(* Logix 5000 project; controller PLC_MCC1300_75F1 vendor 1 type 14 code 166 rev 32.11; software revision 32.04; part 73 of 83 *)
(* tags used below, declared in another part *)
   GP_OB_InitializeMain : GP_OB_Initialize;
   GP_RampSpace : GP_RampSpace;
   GP_ScadaPlate : GP_ScadaPlate;
   Gp_SpaceConvUtilities_V1 : GP_SpaceConvUtilities_V1;
   M351 : MAC_Conveyor;
   M351_Data : UDT_Convoy_SL;
   M351_SpaceConv_Utilities : SpaceConv_Utilities;
   M352 : MAC_Conveyor;
   M352_ALM : MAC_Conveyor_ALM;
   M352_Data : UDT_Convoy_SL;
   M352_DeletePlate : BOOL;
   M352_HMR : MAC_Conveyor_HMR;
   M352_HMW : MAC_Conveyor_HMW;
   M352_Input_xPbDeleteGlass : BOOL;
   M352_Input_xPbFanOff : BOOL;   // W204SB3/A. Fan off
   M352_Input_xPbSendToCullet : BOOL;   // W204SB2. Send to cullet
   M352_M1_DR : AXIS_CIP_DRIVE;
   M352_ONS_SetResetPresence : BOOL;
   M352_SpaceConv_Utilities : SpaceConv_Utilities;
   O : INT[128];
   TMP_dConveyorNumberForZoneCleaning : DINT;
   TMP_dDecelerationPositionEndConveyor : DINT;
   TMP_dOffsetLoadUnload_cmm : DINT;
   TMP_SendToCullet : BOOL;
   TMP_x : BOOL;
   TMP_xConveyorInvolvedInCleaning : BOOL;
   TMP_xConveyorOfStartCleaning : BOOL;
   TMP_xEnableLoadUnload : BOOL;
   TMP_xEnableZoneCleaning : BOOL;
   xAlwaysOFF : BOOL;
   xAlwaysON : BOOL;
   xSampleTablePedal : BOOL;
   Z900 : MAC_Zone;
   Z900_HMI_rgtPlateScada_Internal : HMI_LiteData[5,2,7];
   Z900_HMW : MAC_Zone_HMW;
(* MainProgram, continued *)

ROUTINE M352_Alarm   (* ladder *)
   0: NOP();
   // Reset Alarm
   1: XIC(Z900.tmON_ResetAlarm.DN)FLL(0,M352_ALM,1);
   2: XIC(Z900.ST_xEnableControlError)XIC(xAlwaysOFF)XIO(M352.INPUT_xProtectionMotor_M1)OTL(M352_ALM.rgxStoppingFault_M[0].0);
   3: XIC(Z900.ST_xEnableControlError)XIC(M352.INPUT_xDriveError_M1)OTL(M352_ALM.rgxStoppingFault_M[0].1);
   4: XIC(Z900.ST_xEnableControlError)XIO(M352.INPUT_xDriveError_M1)[XIC(M352.OUTPUT_xRun_M1) ,XIC(M352.OUTPUT_xReverse_M1) ,XIC(M352.OUTPUT_xPositioning_M1) ]XIO(M352.INPUT_xDriveFeedback_M1)[XIO(M352.tmON_FeedbackTimeOut_M1.DN) TON(M352.tmON_FeedbackTimeOut_M1,?,?) ,XIC(M352.tmON_FeedbackTimeOut_M1.DN) OTL(M352_ALM.rgxStoppingFault_M[0].2) ];
   5: XIC(Z900.ST_xEnableControlError)XIC(xAlwaysOFF)XIO(M352.INPUT_xLocalSafetySwitch_M1)OTL(M352_ALM.rgxStoppingFault_M[0].3);
   6: XIC(Z900.ST_xEnableControlError)XIO(M352.INPUT_xMotorThermalProbe_M1)OTL(M352_ALM.rgxStoppingFault_M[0].4);
   7: XIC(Z900.ST_xEnableControlError)XIC(xAlwaysOFF)XIO(M352.INPUT_xBrakingResistor_M1)OTL(M352_ALM.rgxStoppingFault_M[0].5);
   8: XIC(Z900.ST_xEnableControlError)XIC(xAlwaysOFF)[XIC(M352.INPUT_xDriveInhibit_M1) ,XIC(M352.OUTPUT_xDriveEnable_M1) XIO(M352.INPUT_xDriveReady_M1) ]OTL(M352_ALM.rgxStoppingFault_M[0].6);
   9: XIC(M352.ST_xEnableControlError)XIC(xAlwaysOFF)XIC(M352.PH_x.23)NEQ(M352_SpaceConv_Utilities.CONST_dSyncMode,0)[XIO(M352.ST_xPlateSynchronized) OTL(M352_ALM.rgxWarning[0].0) ,XIC(M352.ST_xPlateSynchronized) OTU(M352_ALM.rgxWarning[0].0) ];
   10: XIC(M352.ST_xEnableControlError)XIC(xAlwaysOFF)XIC(M352.PH_x.23)[XIC(M352_Data.tFlag.tConveyor.xReqStop) ,XIC(M352_Data.tFlag.tConveyor.xBypassReqEndStop) ]OTL(M352_ALM.rgxWarning[0].1);
   // #####_CUMULATIVE ALARM_#####
   11: NOP();
   12: [NEQ(M352_ALM.rgxStoppingFault[0],0) ,NEQ(M352_ALM.rgxStoppingFault_M[0],0) ,NEQ(M352_ALM.rgxStoppingFault_M[1],0) ]OTE(M352.ST_xStopMachineFault);
   13: [NEQ(M352_ALM.rgxFault[0],0) ,NEQ(M352_ALM.rgxFault_M[0],0) ,NEQ(M352_ALM.rgxFault_M[1],0) ]OTE(M352.ST_xStopNextCycleFault);
END_ROUTINE

ROUTINE M352_Logic   (* ladder *)
   // #####_COSTANTS_#####
   0: [MOV(6010,TMP_dConveyorNumberForZoneCleaning) MOV(50000,TMP_dOffsetLoadUnload_cmm) MOV(500,M352_SpaceConv_Utilities.CONST_dPresetFeedbackTime_ms) OTU(TMP_xEnableLoadUnload) OTU(TMP_xEnableZoneCleaning) MOV(500000,M352_SpaceConv_Utilities.CONST_dConveyorLength_cmm) MOV(400000,M352_SpaceConv_Utilities.CONST_dConveyorWidth_cmm) SUB(M352_SpaceConv_Utilities.CONST_dConveyorLength_cmm,M352.AUX_dAccSpace_cmm,M352.AUX_dPresetStopLoad_cmm) ADD(M352_SpaceConv_Utilities.CONST_dConveyorLength_cmm,M352.AUX_dDecSpace_cmm,M352.AUX_dPresetStopUnload_cmm) MOV(1.2,M352_SpaceConv_Utilities.CONST_rAcceleration_ms2) MOV(1.2,M352_SpaceConv_Utilities.CONST_rDeceleration_ms2) ,[MOV(1,M352_SpaceConv_Utilities.CONST_dSyncMode) ,MOV(0,M352_SpaceConv_Utilities.CONST_dSyncroPhPosition_cmm) ,MOV(200000,M352_SpaceConv_Utilities.CONST_dSyncroPhWindow_cmm) ] ];
   // #####_MATCH_#####
   1: NOP();
   // Conveyor Cleaning
   2: XIC(TMP_xEnableZoneCleaning)XIC(Z900.ST_xCleaningAccepted)GRT(Z900_HMW.dCleaningSelection,0)[EQU(Z900_HMW.dCleaningSelection,TMP_dConveyorNumberForZoneCleaning) OTE(TMP_xConveyorOfStartCleaning) ,GEQ(Z900_HMW.dCleaningSelection,TMP_dConveyorNumberForZoneCleaning) OTE(TMP_xConveyorInvolvedInCleaning) ];
   // Enable control error
   3: XIC(Z900.ST_xEnableControlError)OTE(M352.ST_xEnableControlError);
   // Mode 7 - Offsett for load/unload Simultaney
   4: XIC(M352.PH_x.8)MOV(M352.AUX_dPresetStopLoad_cmm,M352_SpaceConv_Utilities.ST_dStopLoadForseen_cmm)MOV(TMP_dOffsetLoadUnload_cmm,M352_SpaceConv_Utilities.CONF_MD7_dOffset_cmm)GP_SpaceConvUtilities_V1(Gp_SpaceConvUtilities_V1,M352_SpaceConv_Utilities,M352_SpaceConv_Utilities,M351_SpaceConv_Utilities,7);
   // #####_ALARMS_#####
   5: NOP();
   // Call Alarm Routine
   6: JSR(M352_Alarm,0);
   // #####_HMI_LOGICS_#####
   7: NOP();
   // Condition ok for Cleaning
   8: [XIO(TMP_xEnableZoneCleaning) ,XIC(TMP_xEnableZoneCleaning) [XIC(M352.ST_xOutputEnable) ,XIO(xAlwaysOFF) ] [XIO(TMP_xConveyorOfStartCleaning) ,XIC(M352.PH_x.0) ,XIO(M352.PH_x.8) ] ]OTE(M352.ST_xCleaningConditionOK);
   // Cleaning Accepted
   9: [[XIC(M352_HMW.xStopLocalCleaningRequest) ,XIC(M352_Input_xPbDeleteGlass) XIO(M352.ST_xPlatePresence) ] OTU(M352_HMW.xStopLocalCleaningRequest) OTU(M352_HMW.xLocalCleaningRequest) ,[XIC(M352_HMW.xLocalCleaningRequest) ,XIC(M352_Input_xPbDeleteGlass) XIC(M352.ST_xPlatePresence) ] [XIC(M352.ST_xCleaningConditionOK) ,XIC(M352.ST_xCleaningAccepted) ] OTE(M352.ST_xCleaningAccepted) ];
   // Manual Mode Enabled
   10: XIO(M352_SpaceConv_Utilities.ST_xFeedbackRotation)[XIC(M352_HMW.xEnableDisableManualCommand) XIC(M352.ST_xConditionOKStopCycle) OTL(M352.ST_xManualMode) ,XIO(M352_HMW.xEnableDisableManualCommand) OTU(M352.ST_xManualMode) ];
   // Virtual door enabled
   11: XIC(M352_HMW.xEnableDisableVirtualDoor)OTE(M352.ST_xVirtualDoorEnabled);
   // Clear manual command
   12: XIO(M352.ST_xManualMode)MOV(0,M352_HMW.rgxMan);
   // #####_STATUSES_#####
   13: NOP();
   // Machine in Alarm
   14: [XIC(M352.ST_xStopMachineFault) ,XIC(M352.ST_xStopNextCycleFault) ]OTE(M352.ST_xMachineAlarm);
   // Condition ok for stop Cycle
   15: [XIO(M352.ST_xPhasesInProgress) ,XIC(M352.PH_x.8) XIO(M352.OUTPUT_xRun_M1) XIO(M352_SpaceConv_Utilities.ST_xFeedbackRotation) ,XIC(M352.ST_xMachineAlarm) ,XIO(Z900.ST_xCycleON) ]OTE(M352.ST_xConditionOKStopCycle);
   // Cycle load unload simultaneous
   16: XIC(TMP_xEnableLoadUnload)XIO(M352.ST_xDisableLoadUnloadOnStop)XIO(M352.ST_xIdPlatePresence)OTE(M352.ST_xCycleLoadUnload);
   // Speed Management
   17: [XIO(M352_SpaceConv_Utilities.O_xRampInProgress) XIO(M352.ST_xManualMode) MOV(40000,M352.AUX_dReqSpeed_mm_min) ,XIC(M352.ST_xManualMode) MOV(Z900_HMW.dManualSpeed_mm_min,M352.AUX_dReqSpeed_mm_min) ,NEQ(M352.AUX_dReqSpeed_mm_min,M352_SpaceConv_Utilities.ST_dRealSpeed_mm_min) OTE(M352.OS_xChangeSpeed) ];
   // Ramp Management
   18: GP_RampSpace(GP_RampSpace,M352_SpaceConv_Utilities.CONST_rAcceleration_ms2,M352_SpaceConv_Utilities.CONST_rDeceleration_ms2,M352_SpaceConv_Utilities.ST_dRealSpeed_mm_min,M352.AUX_dAccSpace_cmm,M352.AUX_dDecSpace_cmm);
   // Space Convoy utilities MOD 1 for Calculate Head/Tail
   19: XIC(xAlwaysON)[[XIC(M352.OUTPUT_xRun_M1) ,XIC(M352.OUTPUT_xReverse_M1) ] XIO(M352.ST_xManualMode) OTE(M352_SpaceConv_Utilities.CONF_MD1_xRun) ,XIC(M352.OUTPUT_xReverse_M1) XIC(xAlwaysOFF) XIO(M352.ST_xManualMode) OTE(M352_SpaceConv_Utilities.CONF_MD1_xReverse) ,[XIC(M352.INPUT_xDriveFeedback_M1) ,XIC(M352_SpaceConv_Utilities.CONF_MD1_xRun) GRT(M352_SpaceConv_Utilities.O_dCountFeedbackTime_ms,0) ] OTE(M352_SpaceConv_Utilities.ST_xFeedbackRotation) ,XIC(M352.ST_xIdPlatePresence) OTE(M352_SpaceConv_Utilities.CONF_MD1_xHeadTracking) ,XIC(M352.ST_xPlatePresence) OTE(M352_SpaceConv_Utilities.CONF_MD1_xTailTracking) ,MOV(GP_OB_InitializeMain.OUT_dExecutionTime_ms,M352_SpaceConv_Utilities.CONF_MD1_dScan_ms) GP_SpaceConvUtilities_V1(Gp_SpaceConvUtilities_V1,M352_SpaceConv_Utilities,M352_SpaceConv_Utilities,M352_SpaceConv_Utilities,1) ];
   // Output Enable
   20: XIC(Z900.ST_xCycleON)XIO(M352.ST_xManualMode)XIO(M352.ST_xStopMachineFault)[XIO(M352.ST_xPlatePassageUpstream_FW) XIO(M352.ST_xPlatePassageUpstream_BKW) ,XIC(M352.ST_xPlatePassageUpstream_FW) XIC(xAlwaysOFF) ,XIC(M352.ST_xPlatePassageUpstream_BKW) XIC(M351.ST_xOutputEnable) ]OTE(M352.ST_xOutputEnable);
   // #####_WORKING_FLAGS_#####
   21: NOP();
   // #####_LOGICS_#####
   22: NOP();
   // Phase of load (from M351)
   23: XIC(M351.OS_xUnload_BW)[OTL(M352.PH_x.16) ,OTU(M352_SpaceConv_Utilities.O_xPlateSynchronized) ,OTU(M352.ST_xDisableLoadUnloadOnStop) ,OTE(M352.OS_xLoad_BW) ,COP(M351_Data,M352_Data,1) FLL(0,M351_Data,1) ,GP_SpaceConvUtilities_V1(Gp_SpaceConvUtilities_V1,M352_SpaceConv_Utilities,M352_SpaceConv_Utilities,M351_SpaceConv_Utilities,15) ];
   // End load Phase (from M351)
   24: XIC(M352.PH_x.16)GRT(M352_SpaceConv_Utilities.O_dHeadPosition_cmm,M352.AUX_dPresetStopLoad_cmm)[OTE(M352.PH_x.23) ,OTU(M352.PH_x.16) ,OTL(M352.PH_x.24) ,OTL(M352.ST_xPlatePresence) ];
   25: XIC(M352.PH_x.24)XIC(M352_Input_xPbFanOff)[OTU(M352.PH_x.24) ,OTE(M352_DeletePlate) ];
   // Calculation Space for Wait Stop Next Conveyor
   26: CPT(TMP_dDecelerationPositionEndConveyor,M352_SpaceConv_Utilities.CONST_dConveyorLength_cmm - M352.AUX_dAccSpace_cmm + 1000);
   // Wait stop next Machine
   27: XIO(M352.PH_x.8)GEQ(M352_SpaceConv_Utilities.O_dHeadPosition_cmm,TMP_dDecelerationPositionEndConveyor)OTE(M352.ST_xWaitStopNextMachine);
   28: XIC(xAlwaysON)XIC(xSampleTablePedal)OTE(M352.ST_xAux1);
   // Phase of unload to sample table
   29: XIC(Z900.ST_xConditionOkPhaseAdvancement)XIC(M352.ST_xPlatePresence)XIC(M352.ST_xIdPlatePresence)XIC(M352.ST_xOutputEnable)XIO(M352.ST_xWaitMachineStop)XIO(M352.PH_x.8)[XIC(M352.ST_xAux1) [OTE(M352.ST_xWaitReadyToMove) ,[XIC(M352.ST_xAxleReadyToMoveDelayed) ,XIC(xAlwaysON) ] [OTE(M352.OS_xUnload_FW) ,OTL(M352.PH_x.8) ,MOV(M352_Data.dLength_cmm,M352_SpaceConv_Utilities.CONF_MD4_MD6_dLength_cmm) GP_SpaceConvUtilities_V1(Gp_SpaceConvUtilities_V1,M352_SpaceConv_Utilities,M351_SpaceConv_Utilities,M352_SpaceConv_Utilities,6) ] ] ,OTE(M352.ST_xAux2) ];
   // Phase of end unload
   30: XIC(M352.PH_x.8)[XIC(xAlwaysOFF) [GEQ(M352_SpaceConv_Utilities.O_dTailPosition_cmm,M352.AUX_dPresetStopUnload_cmm) ,XIO(M352_SpaceConv_Utilities.ST_xFeedbackRotation) GEQ(M352_SpaceConv_Utilities.O_dTailPosition_cmm,M352_SpaceConv_Utilities.CONST_dConveyorLength_cmm) ] ,XIC(M351.PH_x.7) ][OTE(M352.PH_x.15) ,OTU(M352.PH_x.8) ,OTU(M352.ST_xPlatePresence) ];
   31: XIC(M352_Input_xPbFanOff)ONS(M352_ONS_SetResetPresence)XIO(M352.ST_xPhasesInProgress)[XIC(M352.ST_xPlatePresence) OTU(M352.ST_xPlatePresence) OTE(TMP_x) ,XIO(M352.ST_xPlatePresence) XIO(TMP_x) OTL(M352.ST_xPlatePresence) ];
   // Redestination lites
   32: [XIC(M352_Input_xPbSendToCullet) ,XIC(M352_DeletePlate) ]OTE(TMP_SendToCullet)XIC(M352_DeletePlate)OTU(M352.ST_xPlatePresence)FLL(0,M352_Data,1);
   // Phase in progress
   33: NEQ(M352.PH_x,0)OTE(M352.ST_xPhasesInProgress);
   // #####_CLEANING_#####
   34: NOP();
   // Cleaning Reset
   35: XIC(M352.ST_xCleaningAccepted)[XIC(Z900.ST_xCleaningAccepted) ,XIO(TMP_xConveyorOfStartCleaning) ][XIC(M352.ST_xIdPlatePresence) OTL(TMP_SendToCullet) FLL(0,M352_Data,1) ,MOV(0,M352.PH_x) OTU(M352.ST_xPlatePresence) ];
   // Initial condition OK
   36: XIC(Z900.ST_xConditionOkPhaseAdvancement)XIC(M352.ST_xOutputEnable)XIO(M352_HMW.xEnableDisableManualCommand)XIO(M352.ST_xReqCleaning)XIO(M352.ST_xCleaningAccepted)XIO(M352.ST_xStopNextCycleFault)XIO(M352.ST_xVirtualDoorEnabled)XIO(M352.PH_x.16)[XIO(M352.ST_xPhasesInProgress) XIO(M352.ST_xPlatePresence) ,XIO(xAlwaysOFF) XIC(M352.ST_xCycleLoadUnload) XIC(M352.PH_x.8) XIC(M352.OUTPUT_xRun_M1) GRT(M352_SpaceConv_Utilities.O_dTailPosition_cmm,M352_SpaceConv_Utilities.O_dPresetLoadUnload_cmm) XIO(M352.ST_xIdPlatePresence) ][XIC(M352.INPUT_xHighPositionPopup_1) XIC(M352.ST_xAux1) OTE(M352.ST_xInitialConditionOK) ,OTE(M352.ST_xAux3) ];
   // #####_HMI_STATUSES_#####
   37: NOP();
   // Manual Mode Enable {x|x|x|x|O}
   38: XIC(M352.ST_xManualMode)OTE(M352_HMR.xManualCommandEnabled);
   // Command forward M1
   39: XIC(M352.ST_xManualMode)XIC(M352_HMW.rgxMan.0)XIC(M352.OUTPUT_xRun_M1)OTE(M352_HMR.rgxMan.0);
   // Command backward M1
   40: XIC(M352.ST_xManualMode)XIC(M352_HMW.rgxMan.1)XIC(M352.OUTPUT_xReverse_M1)OTE(M352_HMR.rgxMan.1);
   // Command M2 start air cushion
   41: XIC(M352.ST_xManualMode)XIC(M352_HMW.rgxMan.14)XIC(M352.OUTPUT_xRun_M2)OTE(M352_HMR.rgxMan.14);
   // Command M2 stop air cushion
   42: XIC(M352.ST_xManualMode)XIC(M352_HMW.rgxMan.15)XIO(M352.OUTPUT_xRun_M2)OTE(M352_HMR.rgxMan.15);
   // Cleaning Enabled {x|x|x|x|O}
   43: XIC(M352.ST_xCleaningAccepted)[XIC(Z900.ST_xCleaningAccepted) ,XIO(TMP_xEnableZoneCleaning) ,]OTE(M352_HMR.xCleaningEnabled);
   // Virtual door Enabled {x|x|x|x|O}
   44: XIC(M352.ST_xVirtualDoorEnabled)OTE(M352_HMR.xVirtualDoorEnabled);
   // Id plate presence
   45: XIC(M352.ST_xIdPlatePresence)OTE(M352_HMR.xIdPlatePresence);
   // Machine state M1
   46: XIC(xAlwaysON)[MOV(1,M352_HMR.dState1) ,XIC(M352.OUTPUT_xRun_M1) MOV(3,M352_HMR.dState1) ,XIC(M352.OUTPUT_xReverse_M1) MOV(4,M352_HMR.dState1) ,XIC(M352.ST_xMachineAlarm) MOV(7,M352_HMR.dState1) ];
   // Machine state M2
   47: XIC(xAlwaysON)[MOV(1,M352_HMR.dState2) ,XIC(M352.OUTPUT_xRun_M2) MOV(3,M352_HMR.dState2) ,XIC(M352.OUTPUT_xReverse_M2) MOV(4,M352_HMR.dState2) ,XIC(M352.ST_xMachineAlarm) MOV(7,M352_HMR.dState2) ];
   48: XIC(M352_SpaceConv_Utilities.O_xPlateSynchronized)OTE(M352.ST_xPlateSynchronized);
   // Motor error code
   49: MOV(M352_M1_DR.AxisFault,M352_HMR.dErrorCode1);
   50: XIC(M352.ST_xIdPlatePresence)GP_ScadaPlate(GP_ScadaPlate,M352_Data,1,M352_SpaceConv_Utilities.O_dHeadPosition_cmm,M352_SpaceConv_Utilities.CONST_dConveyorWidth_cmm,M352_SpaceConv_Utilities.CONST_dConveyorLength_cmm,M352_SpaceConv_Utilities.ST_xLastModLoadBkw,M352_SpaceConv_Utilities.ST_xLastModUnloadBkw,1,1,Z900_HMI_rgtPlateScada_Internal);
END_ROUTINE
